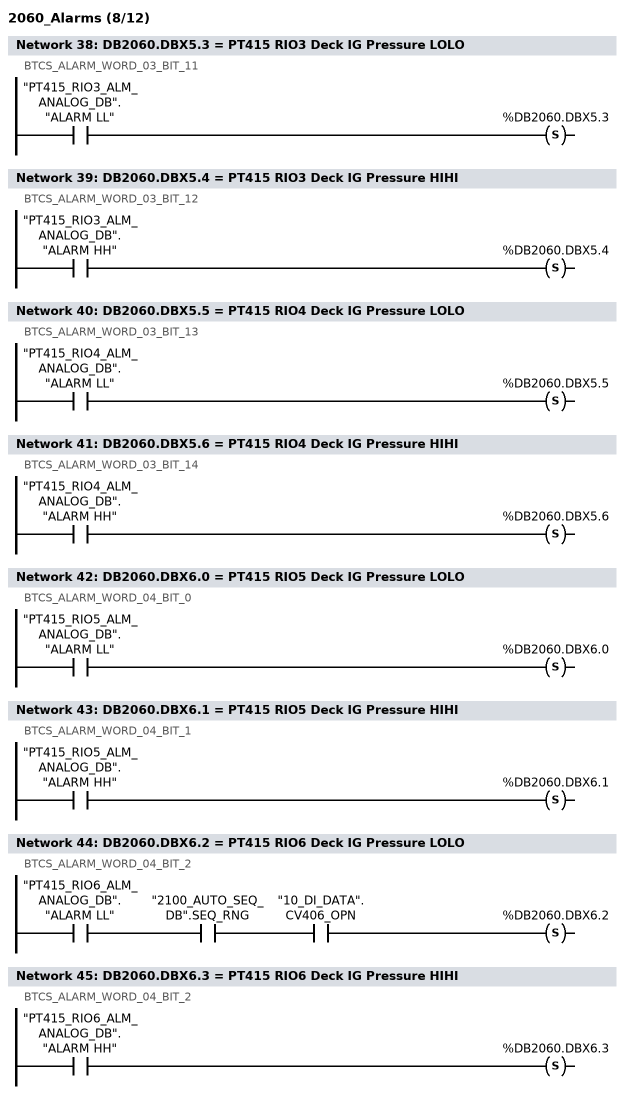
   RUNG wire#powerrail
      Contact( "PT415_RIO3_ALM_ANALOG_DB"."ALARM LL" )
      S_Coil( %DB2060.DBX5.3 )
   END_RUNG
   // the same network as SCL:
   IF "PT415_RIO3_ALM_ANALOG_DB"."ALARM LL" THEN %DB2060.DBX5.3 := TRUE; END_IF;
END_REGION

REGION Network 39: DB2060.DBX5.4 = PT415 RIO3 Deck IG Pressure HIHI
   // BTCS_ALARM_WORD_03_BIT_12
   RUNG wire#powerrail
      Contact( "PT415_RIO3_ALM_ANALOG_DB"."ALARM HH" )
      S_Coil( %DB2060.DBX5.4 )
   END_RUNG
   // the same network as SCL:
   IF "PT415_RIO3_ALM_ANALOG_DB"."ALARM HH" THEN %DB2060.DBX5.4 := TRUE; END_IF;
END_REGION

REGION Network 40: DB2060.DBX5.5 = PT415 RIO4 Deck IG Pressure LOLO
   // BTCS_ALARM_WORD_03_BIT_13
   RUNG wire#powerrail
      Contact( "PT415_RIO4_ALM_ANALOG_DB"."ALARM LL" )
      S_Coil( %DB2060.DBX5.5 )
   END_RUNG
   // the same network as SCL:
   IF "PT415_RIO4_ALM_ANALOG_DB"."ALARM LL" THEN %DB2060.DBX5.5 := TRUE; END_IF;
END_REGION

REGION Network 41: DB2060.DBX5.6 = PT415 RIO4 Deck IG Pressure HIHI
   // BTCS_ALARM_WORD_03_BIT_14
   RUNG wire#powerrail
      Contact( "PT415_RIO4_ALM_ANALOG_DB"."ALARM HH" )
      S_Coil( %DB2060.DBX5.6 )
   END_RUNG
   // the same network as SCL:
   IF "PT415_RIO4_ALM_ANALOG_DB"."ALARM HH" THEN %DB2060.DBX5.6 := TRUE; END_IF;
END_REGION

REGION Network 42: DB2060.DBX6.0 = PT415 RIO5 Deck IG Pressure LOLO
   // BTCS_ALARM_WORD_04_BIT_0
   RUNG wire#powerrail
      Contact( "PT415_RIO5_ALM_ANALOG_DB"."ALARM LL" )
      S_Coil( %DB2060.DBX6.0 )
   END_RUNG
   // the same network as SCL:
   IF "PT415_RIO5_ALM_ANALOG_DB"."ALARM LL" THEN %DB2060.DBX6.0 := TRUE; END_IF;
END_REGION

REGION Network 43: DB2060.DBX6.1 = PT415 RIO5 Deck IG Pressure HIHI
   // BTCS_ALARM_WORD_04_BIT_1
   RUNG wire#powerrail
      Contact( "PT415_RIO5_ALM_ANALOG_DB"."ALARM HH" )
      S_Coil( %DB2060.DBX6.1 )
   END_RUNG
   // the same network as SCL:
   IF "PT415_RIO5_ALM_ANALOG_DB"."ALARM HH" THEN %DB2060.DBX6.1 := TRUE; END_IF;
END_REGION

REGION Network 44: DB2060.DBX6.2 = PT415 RIO6 Deck IG Pressure LOLO
   // BTCS_ALARM_WORD_04_BIT_2
   RUNG wire#powerrail
      Contact( "PT415_RIO6_ALM_ANALOG_DB"."ALARM LL" )
      Contact( "2100_AUTO_SEQ_DB".SEQ_RNG )
      Contact( "10_DI_DATA".CV406_OPN )
      S_Coil( %DB2060.DBX6.2 )
   END_RUNG
   // the same network as SCL:
   IF "PT415_RIO6_ALM_ANALOG_DB"."ALARM LL" AND "2100_AUTO_SEQ_DB".SEQ_RNG AND "10_DI_DATA".CV406_OPN THEN
       %DB2060.DBX6.2 := TRUE;
   END_IF;
END_REGION

REGION Network 45: DB2060.DBX6.3 = PT415 RIO6 Deck IG Pressure HIHI
   // BTCS_ALARM_WORD_04_BIT_2
   RUNG wire#powerrail
      Contact( "PT415_RIO6_ALM_ANALOG_DB"."ALARM HH" )
      S_Coil( %DB2060.DBX6.3 )
   END_RUNG
   // the same network as SCL:
   IF "PT415_RIO6_ALM_ANALOG_DB"."ALARM HH" THEN %DB2060.DBX6.3 := TRUE; END_IF;
END_REGION

REGION Network 46: DB2060.DBX6.4 = PT415 RIO7 Deck IG Pressure LOLO
   // BTCS_ALARM_WORD_04_BIT_4
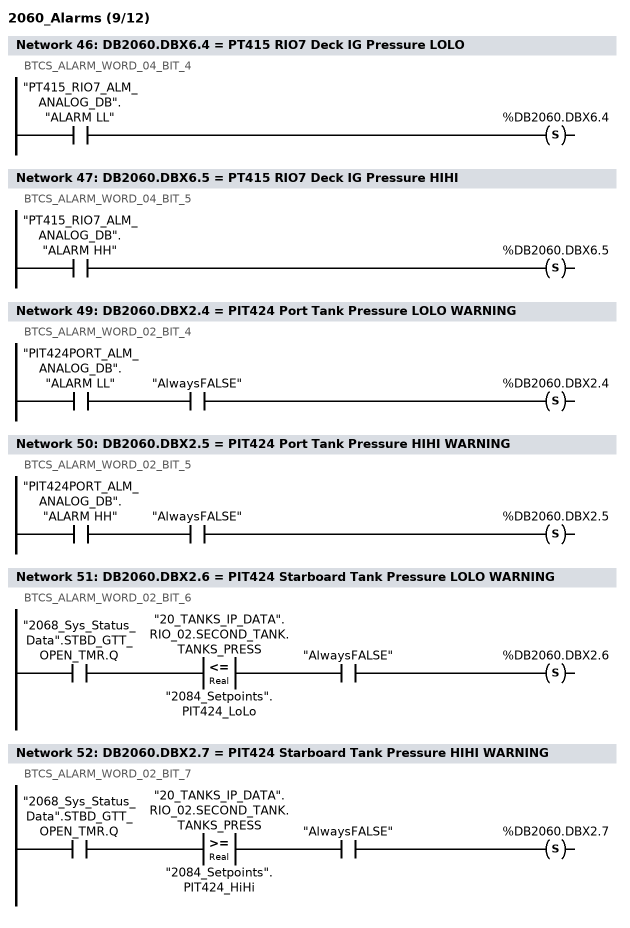
   RUNG wire#powerrail
      Contact( "PT415_RIO7_ALM_ANALOG_DB"."ALARM LL" )
      S_Coil( %DB2060.DBX6.4 )
   END_RUNG
   // the same network as SCL:
   IF "PT415_RIO7_ALM_ANALOG_DB"."ALARM LL" THEN %DB2060.DBX6.4 := TRUE; END_IF;
END_REGION

REGION Network 47: DB2060.DBX6.5 = PT415 RIO7 Deck IG Pressure HIHI
   // BTCS_ALARM_WORD_04_BIT_5
   RUNG wire#powerrail
      Contact( "PT415_RIO7_ALM_ANALOG_DB"."ALARM HH" )
      S_Coil( %DB2060.DBX6.5 )
   END_RUNG
   // the same network as SCL:
   IF "PT415_RIO7_ALM_ANALOG_DB"."ALARM HH" THEN %DB2060.DBX6.5 := TRUE; END_IF;
END_REGION

REGION Network 49: DB2060.DBX2.4 = PIT424 Port Tank Pressure LOLO WARNING
   // BTCS_ALARM_WORD_02_BIT_4
   RUNG wire#powerrail
      Contact( "PIT424PORT_ALM_ANALOG_DB"."ALARM LL" )
      Contact( "AlwaysFALSE" )
      S_Coil( %DB2060.DBX2.4 )
   END_RUNG
   // the same network as SCL:
   IF "PIT424PORT_ALM_ANALOG_DB"."ALARM LL" AND "AlwaysFALSE" THEN %DB2060.DBX2.4 := TRUE; END_IF;
END_REGION

REGION Network 50: DB2060.DBX2.5 = PIT424 Port Tank Pressure HIHI WARNING
   // BTCS_ALARM_WORD_02_BIT_5
   RUNG wire#powerrail
      Contact( "PIT424PORT_ALM_ANALOG_DB"."ALARM HH" )
      Contact( "AlwaysFALSE" )
      S_Coil( %DB2060.DBX2.5 )
   END_RUNG
   // the same network as SCL:
   IF "PIT424PORT_ALM_ANALOG_DB"."ALARM HH" AND "AlwaysFALSE" THEN %DB2060.DBX2.5 := TRUE; END_IF;
END_REGION

REGION Network 51: DB2060.DBX2.6 = PIT424 Starboard Tank Pressure LOLO WARNING
   // BTCS_ALARM_WORD_02_BIT_6
   RUNG wire#powerrail
      Contact( "2068_Sys_Status_Data".STBD_GTT_OPEN_TMR.Q )
      { S7_Templates := "SrcType := Real" } LE_Contact(in1 := "20_TANKS_IP_DATA".RIO_02.SECOND_TANK.TANKS_PRESS, in2 := "2084_Setpoints".PIT424_LoLo)
      Contact( "AlwaysFALSE" )
      S_Coil( %DB2060.DBX2.6 )
   END_RUNG
   // the same network as SCL:
   IF "2068_Sys_Status_Data".STBD_GTT_OPEN_TMR.Q AND ("20_TANKS_IP_DATA".RIO_02.SECOND_TANK.TANKS_PRESS <= "2084_Setpoints".PIT424_LoLo) AND "AlwaysFALSE" THEN
       %DB2060.DBX2.6 := TRUE;
   END_IF;
END_REGION

REGION Network 52: DB2060.DBX2.7 = PIT424 Starboard Tank Pressure HIHI WARNING
   // BTCS_ALARM_WORD_02_BIT_7
   RUNG wire#powerrail
      Contact( "2068_Sys_Status_Data".STBD_GTT_OPEN_TMR.Q )
      { S7_Templates := "SrcType := Real" } GE_Contact(in1 := "20_TANKS_IP_DATA".RIO_02.SECOND_TANK.TANKS_PRESS, in2 := "2084_Setpoints".PIT424_HiHi)
      Contact( "AlwaysFALSE" )
      S_Coil( %DB2060.DBX2.7 )
   END_RUNG
   // the same network as SCL:
   IF "2068_Sys_Status_Data".STBD_GTT_OPEN_TMR.Q AND ("20_TANKS_IP_DATA".RIO_02.SECOND_TANK.TANKS_PRESS >= "2084_Setpoints".PIT424_HiHi) AND "AlwaysFALSE" THEN
       %DB2060.DBX2.7 := TRUE;
   END_IF;
END_REGION

REGION Network 54: Alarm reset
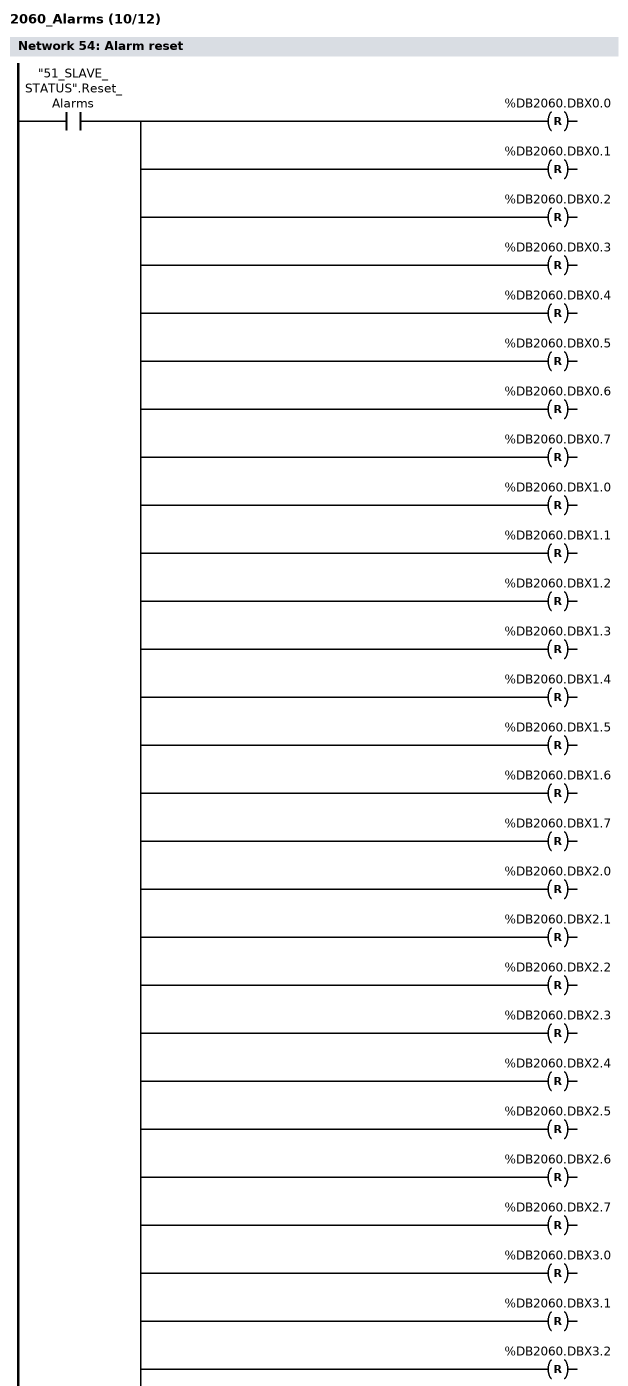
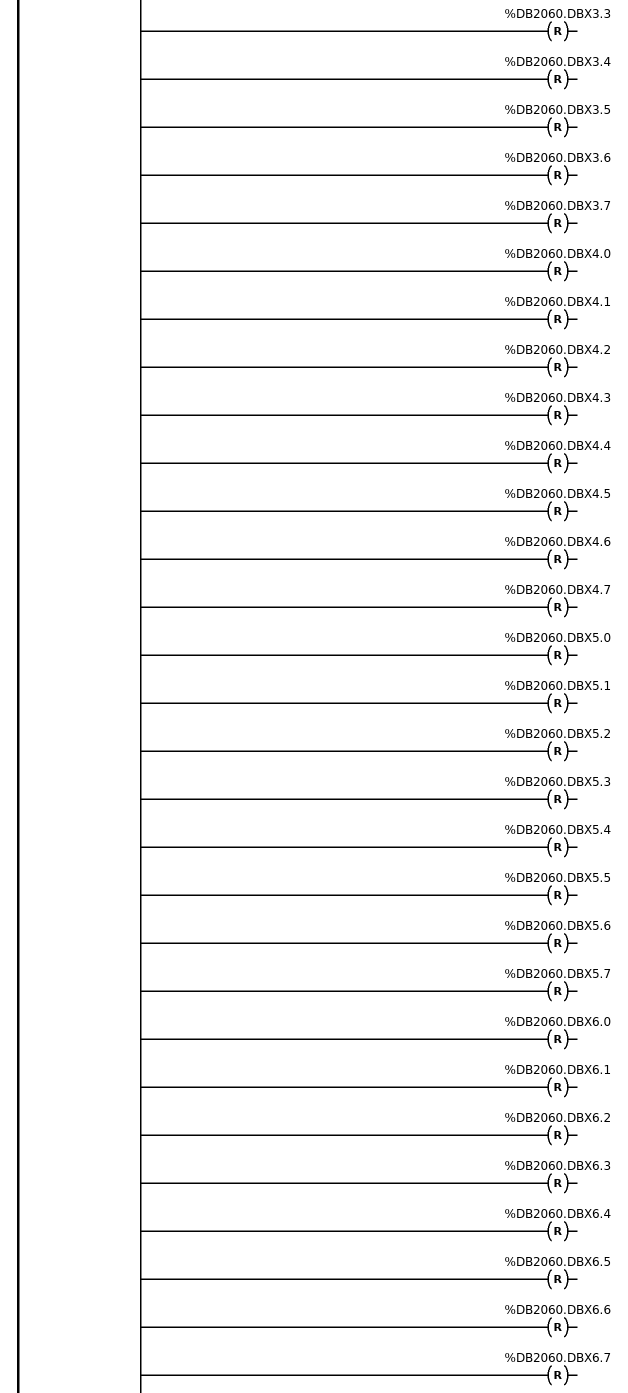
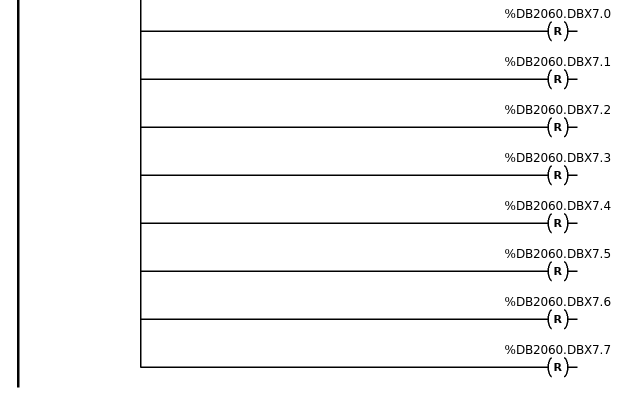
   RUNG wire#powerrail
      Contact( "51_SLAVE_STATUS".Reset_Alarms )
      wire#w1
      R_Coil( %DB2060.DBX0.0 )
   END_RUNG
   RUNG wire#w1
      R_Coil( %DB2060.DBX0.1 )
   END_RUNG
   RUNG wire#w1
      R_Coil( %DB2060.DBX0.2 )
   END_RUNG
   RUNG wire#w1
      R_Coil( %DB2060.DBX0.3 )
   END_RUNG
   RUNG wire#w1
      R_Coil( %DB2060.DBX0.4 )
   END_RUNG
   RUNG wire#w1
      R_Coil( %DB2060.DBX0.5 )
   END_RUNG
   RUNG wire#w1
      R_Coil( %DB2060.DBX0.6 )
   END_RUNG
   RUNG wire#w1
      R_Coil( %DB2060.DBX0.7 )
   END_RUNG
   RUNG wire#w1
      R_Coil( %DB2060.DBX1.0 )
   END_RUNG
   RUNG wire#w1
      R_Coil( %DB2060.DBX1.1 )
   END_RUNG
   RUNG wire#w1
      R_Coil( %DB2060.DBX1.2 )
   END_RUNG
   RUNG wire#w1
      R_Coil( %DB2060.DBX1.3 )
   END_RUNG
   RUNG wire#w1
      R_Coil( %DB2060.DBX1.4 )
   END_RUNG
   RUNG wire#w1
      R_Coil( %DB2060.DBX1.5 )
   END_RUNG
   RUNG wire#w1
      R_Coil( %DB2060.DBX1.6 )
   END_RUNG
   RUNG wire#w1
      R_Coil( %DB2060.DBX1.7 )
   END_RUNG
   RUNG wire#w1
      R_Coil( %DB2060.DBX2.0 )
   END_RUNG
   RUNG wire#w1
      R_Coil( %DB2060.DBX2.1 )
   END_RUNG
   RUNG wire#w1
      R_Coil( %DB2060.DBX2.2 )
   END_RUNG
   RUNG wire#w1
      R_Coil( %DB2060.DBX2.3 )
   END_RUNG
   RUNG wire#w1
      R_Coil( %DB2060.DBX2.4 )
   END_RUNG
   RUNG wire#w1
      R_Coil( %DB2060.DBX2.5 )
   END_RUNG
   RUNG wire#w1
      R_Coil( %DB2060.DBX2.6 )
   END_RUNG
   RUNG wire#w1
      R_Coil( %DB2060.DBX2.7 )
   END_RUNG
   RUNG wire#w1
      R_Coil( %DB2060.DBX3.0 )
   END_RUNG
   RUNG wire#w1
      R_Coil( %DB2060.DBX3.1 )
   END_RUNG
   RUNG wire#w1
      R_Coil( %DB2060.DBX3.2 )
   END_RUNG
   RUNG wire#w1
      R_Coil( %DB2060.DBX3.3 )
   END_RUNG
   RUNG wire#w1
      R_Coil( %DB2060.DBX3.4 )
   END_RUNG
   RUNG wire#w1
      R_Coil( %DB2060.DBX3.5 )
   END_RUNG
   RUNG wire#w1
      R_Coil( %DB2060.DBX3.6 )
   END_RUNG
   RUNG wire#w1
      R_Coil( %DB2060.DBX3.7 )
   END_RUNG
   RUNG wire#w1
      R_Coil( %DB2060.DBX4.0 )
   END_RUNG
   RUNG wire#w1
      R_Coil( %DB2060.DBX4.1 )
   END_RUNG
   RUNG wire#w1
      R_Coil( %DB2060.DBX4.2 )
   END_RUNG
   RUNG wire#w1
      R_Coil( %DB2060.DBX4.3 )
   END_RUNG
   RUNG wire#w1
      R_Coil( %DB2060.DBX4.4 )
   END_RUNG
   RUNG wire#w1
      R_Coil( %DB2060.DBX4.5 )
   END_RUNG
   RUNG wire#w1
      R_Coil( %DB2060.DBX4.6 )
   END_RUNG
   RUNG wire#w1
      R_Coil( %DB2060.DBX4.7 )
   END_RUNG
   RUNG wire#w1
      R_Coil( %DB2060.DBX5.0 )
   END_RUNG
   RUNG wire#w1
      R_Coil( %DB2060.DBX5.1 )
   END_RUNG
   RUNG wire#w1
      R_Coil( %DB2060.DBX5.2 )
   END_RUNG
   RUNG wire#w1
      R_Coil( %DB2060.DBX5.3 )
   END_RUNG
   RUNG wire#w1
      R_Coil( %DB2060.DBX5.4 )
   END_RUNG
   RUNG wire#w1
      R_Coil( %DB2060.DBX5.5 )
   END_RUNG
   RUNG wire#w1
      R_Coil( %DB2060.DBX5.6 )
   END_RUNG
   RUNG wire#w1
      R_Coil( %DB2060.DBX5.7 )
   END_RUNG
   RUNG wire#w1
      R_Coil( %DB2060.DBX6.0 )
   END_RUNG
   RUNG wire#w1
      R_Coil( %DB2060.DBX6.1 )
   END_RUNG
   RUNG wire#w1
      R_Coil( %DB2060.DBX6.2 )
   END_RUNG
   RUNG wire#w1
      R_Coil( %DB2060.DBX6.3 )
   END_RUNG
   RUNG wire#w1
      R_Coil( %DB2060.DBX6.4 )
   END_RUNG
   RUNG wire#w1
      R_Coil( %DB2060.DBX6.5 )
   END_RUNG
   RUNG wire#w1
      R_Coil( %DB2060.DBX6.6 )
   END_RUNG
   RUNG wire#w1
      R_Coil( %DB2060.DBX6.7 )
   END_RUNG
   RUNG wire#w1
      R_Coil( %DB2060.DBX7.0 )
   END_RUNG
   RUNG wire#w1
      R_Coil( %DB2060.DBX7.1 )
   END_RUNG
   RUNG wire#w1
      R_Coil( %DB2060.DBX7.2 )
   END_RUNG
   RUNG wire#w1
      R_Coil( %DB2060.DBX7.3 )
   END_RUNG
   RUNG wire#w1
      R_Coil( %DB2060.DBX7.4 )
   END_RUNG
   RUNG wire#w1
      R_Coil( %DB2060.DBX7.5 )
   END_RUNG
   RUNG wire#w1
      R_Coil( %DB2060.DBX7.6 )
   END_RUNG
   RUNG wire#w1
      R_Coil( %DB2060.DBX7.7 )
   END_RUNG
   // the same network as SCL:
   IF "51_SLAVE_STATUS".Reset_Alarms THEN
       %DB2060.DBX0.0 := FALSE;
       %DB2060.DBX0.1 := FALSE;
       %DB2060.DBX0.2 := FALSE;
       %DB2060.DBX0.3 := FALSE;
       %DB2060.DBX0.4 := FALSE;
       %DB2060.DBX0.5 := FALSE;
       %DB2060.DBX0.6 := FALSE;
       %DB2060.DBX0.7 := FALSE;
       %DB2060.DBX1.0 := FALSE;
       %DB2060.DBX1.1 := FALSE;
       %DB2060.DBX1.2 := FALSE;
       %DB2060.DBX1.3 := FALSE;
       %DB2060.DBX1.4 := FALSE;
       %DB2060.DBX1.5 := FALSE;
       %DB2060.DBX1.6 := FALSE;
       %DB2060.DBX1.7 := FALSE;
       %DB2060.DBX2.0 := FALSE;
       %DB2060.DBX2.1 := FALSE;
       %DB2060.DBX2.2 := FALSE;
       %DB2060.DBX2.3 := FALSE;
       %DB2060.DBX2.4 := FALSE;
       %DB2060.DBX2.5 := FALSE;
       %DB2060.DBX2.6 := FALSE;
       %DB2060.DBX2.7 := FALSE;
       %DB2060.DBX3.0 := FALSE;
       %DB2060.DBX3.1 := FALSE;
       %DB2060.DBX3.2 := FALSE;
       %DB2060.DBX3.3 := FALSE;
       %DB2060.DBX3.4 := FALSE;
       %DB2060.DBX3.5 := FALSE;
       %DB2060.DBX3.6 := FALSE;
       %DB2060.DBX3.7 := FALSE;
       %DB2060.DBX4.0 := FALSE;
       %DB2060.DBX4.1 := FALSE;
       %DB2060.DBX4.2 := FALSE;
       %DB2060.DBX4.3 := FALSE;
       %DB2060.DBX4.4 := FALSE;
       %DB2060.DBX4.5 := FALSE;
       %DB2060.DBX4.6 := FALSE;
       %DB2060.DBX4.7 := FALSE;
       %DB2060.DBX5.0 := FALSE;
       %DB2060.DBX5.1 := FALSE;
       %DB2060.DBX5.2 := FALSE;
       %DB2060.DBX5.3 := FALSE;
       %DB2060.DBX5.4 := FALSE;
       %DB2060.DBX5.5 := FALSE;
       %DB2060.DBX5.6 := FALSE;
       %DB2060.DBX5.7 := FALSE;
       %DB2060.DBX6.0 := FALSE;
       %DB2060.DBX6.1 := FALSE;
       %DB2060.DBX6.2 := FALSE;
       %DB2060.DBX6.3 := FALSE;
       %DB2060.DBX6.4 := FALSE;
       %DB2060.DBX6.5 := FALSE;
       %DB2060.DBX6.6 := FALSE;
       %DB2060.DBX6.7 := FALSE;
       %DB2060.DBX7.0 := FALSE;
       %DB2060.DBX7.1 := FALSE;
       %DB2060.DBX7.2 := FALSE;
       %DB2060.DBX7.3 := FALSE;
       %DB2060.DBX7.4 := FALSE;
       %DB2060.DBX7.5 := FALSE;
       %DB2060.DBX7.6 := FALSE;
       %DB2060.DBX7.7 := FALSE;
   END_IF;
END_REGION

REGION Network 55: New Alarm
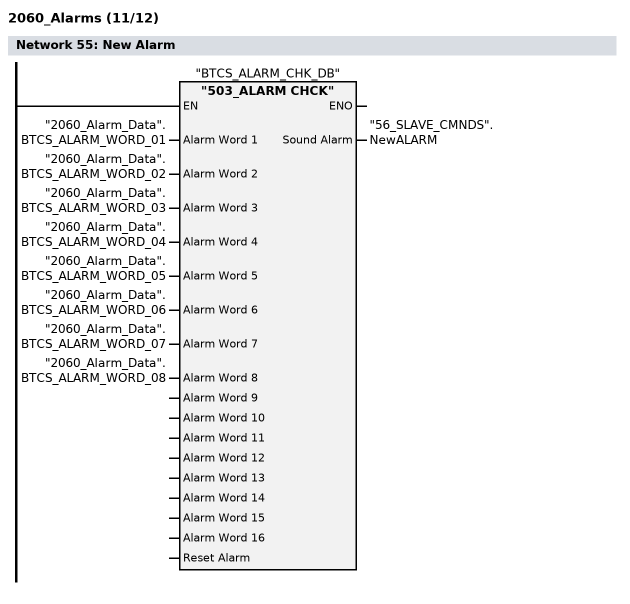
   RUNG wire#powerrail
      "BTCS_ALARM_CHK_DB"("Alarm Word 1" := "2060_Alarm_Data".BTCS_ALARM_WORD_01, "Alarm Word 2" := "2060_Alarm_Data".BTCS_ALARM_WORD_02, "Alarm Word 3" := "2060_Alarm_Data".BTCS_ALARM_WORD_03, "Alarm Word 4" := "2060_Alarm_Data".BTCS_ALARM_WORD_04, "Alarm Word 5" := "2060_Alarm_Data".BTCS_ALARM_WORD_05, "Alarm Word 6" := "2060_Alarm_Data".BTCS_ALARM_WORD_06, "Alarm Word 7" := "2060_Alarm_Data".BTCS_ALARM_WORD_07, "Alarm Word 8" := "2060_Alarm_Data".BTCS_ALARM_WORD_08, "Alarm Word 9" :=, "Alarm Word 10" :=, "Alarm Word 11" :=, "Alarm Word 12" :=, "Alarm Word 13" :=, "Alarm Word 14" :=, "Alarm Word 15" :=, "Alarm Word 16" :=, "Reset Alarm" :=, "Sound Alarm" => "56_SLAVE_CMNDS".NewALARM)
   END_RUNG
   // the same network as SCL:
   "BTCS_ALARM_CHK_DB"("Alarm Word 1" := "2060_Alarm_Data".BTCS_ALARM_WORD_01,   // "503_ALARM CHCK"
                       "Alarm Word 2" := "2060_Alarm_Data".BTCS_ALARM_WORD_02,
                       "Alarm Word 3" := "2060_Alarm_Data".BTCS_ALARM_WORD_03,
                       "Alarm Word 4" := "2060_Alarm_Data".BTCS_ALARM_WORD_04,
                       "Alarm Word 5" := "2060_Alarm_Data".BTCS_ALARM_WORD_05,
                       "Alarm Word 6" := "2060_Alarm_Data".BTCS_ALARM_WORD_06,
                       "Alarm Word 7" := "2060_Alarm_Data".BTCS_ALARM_WORD_07,
                       "Alarm Word 8" := "2060_Alarm_Data".BTCS_ALARM_WORD_08,
                       "Sound Alarm" => "56_SLAVE_CMNDS".NewALARM);
END_REGION

REGION Network 56: Alarm Present
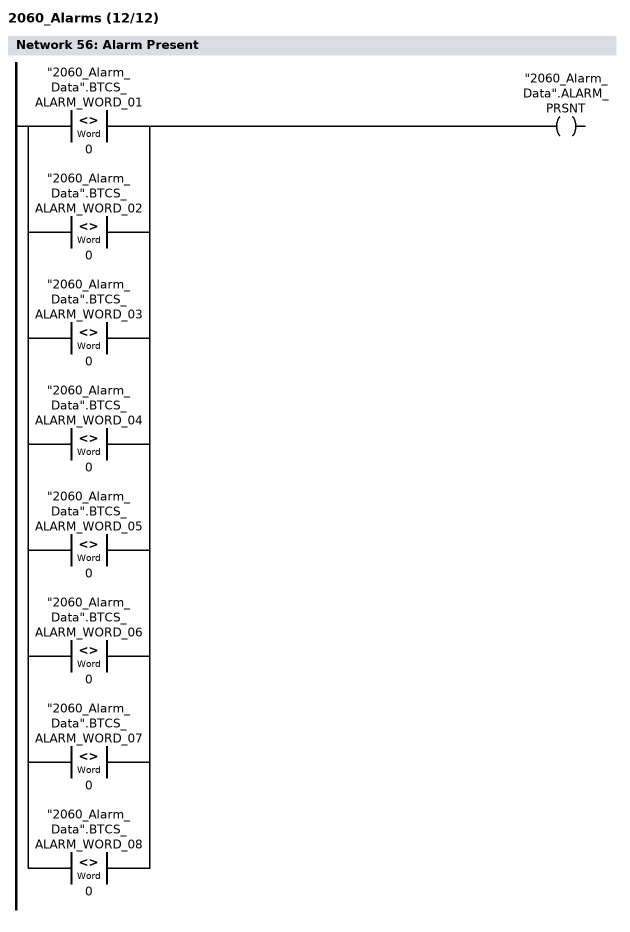
   RUNG wire#powerrail
      { S7_Templates := "SrcType := Word" } NE_Contact(in1 := "2060_Alarm_Data".BTCS_ALARM_WORD_01, in2 := 0)
      wire#w1
      Coil( "2060_Alarm_Data".ALARM_PRSNT )
   END_RUNG
   RUNG wire#powerrail
      { S7_Templates := "SrcType := Word" } NE_Contact(in1 := "2060_Alarm_Data".BTCS_ALARM_WORD_02, in2 := 0)
   END_RUNG wire#w1
   RUNG wire#powerrail
      { S7_Templates := "SrcType := Word" } NE_Contact(in1 := "2060_Alarm_Data".BTCS_ALARM_WORD_03, in2 := 0)
   END_RUNG wire#w1
   RUNG wire#powerrail
      { S7_Templates := "SrcType := Word" } NE_Contact(in1 := "2060_Alarm_Data".BTCS_ALARM_WORD_04, in2 := 0)
   END_RUNG wire#w1
   RUNG wire#powerrail
      { S7_Templates := "SrcType := Word" } NE_Contact(in1 := "2060_Alarm_Data".BTCS_ALARM_WORD_05, in2 := 0)
   END_RUNG wire#w1
   RUNG wire#powerrail
      { S7_Templates := "SrcType := Word" } NE_Contact(in1 := "2060_Alarm_Data".BTCS_ALARM_WORD_06, in2 := 0)
   END_RUNG wire#w1
   RUNG wire#powerrail
      { S7_Templates := "SrcType := Word" } NE_Contact(in1 := "2060_Alarm_Data".BTCS_ALARM_WORD_07, in2 := 0)
   END_RUNG wire#w1
   RUNG wire#powerrail
      { S7_Templates := "SrcType := Word" } NE_Contact(in1 := "2060_Alarm_Data".BTCS_ALARM_WORD_08, in2 := 0)
   END_RUNG wire#w1
   // the same network as SCL:
   "2060_Alarm_Data".ALARM_PRSNT := ("2060_Alarm_Data".BTCS_ALARM_WORD_01 <> 0) OR ("2060_Alarm_Data".BTCS_ALARM_WORD_02 <> 0) OR ("2060_Alarm_Data".BTCS_ALARM_WORD_03 <> 0) OR ("2060_Alarm_Data".BTCS_ALARM_WORD_04 <> 0) OR ("2060_Alarm_Data".BTCS_ALARM_WORD_05 <> 0) OR ("2060_Alarm_Data".BTCS_ALARM_WORD_06 <> 0) OR ("2060_Alarm_Data".BTCS_ALARM_WORD_07 <> 0) OR ("2060_Alarm_Data".BTCS_ALARM_WORD_08 <> 0);
END_REGION
END_FUNCTION

FUNCTION "2062_Warnings" : Void   // FC2062, LAD
TITLE = Warning Processing
{ S7_Optimized_Access := 'TRUE' }
AUTHOR : JRS
VERSION : 0.1
// To warning conditions
   VAR_TEMP   // added for the SCL form of the ladder/FBD networks
      _w1 : Bool;
   END_VAR
BEGIN

REGION Network 1: DB2062 DBX0.0 = 600-TX-433 RIO7 Confined Space O2 Monitor
   // BTCS_WARNING_WORD_01_BIT_0                           15.10
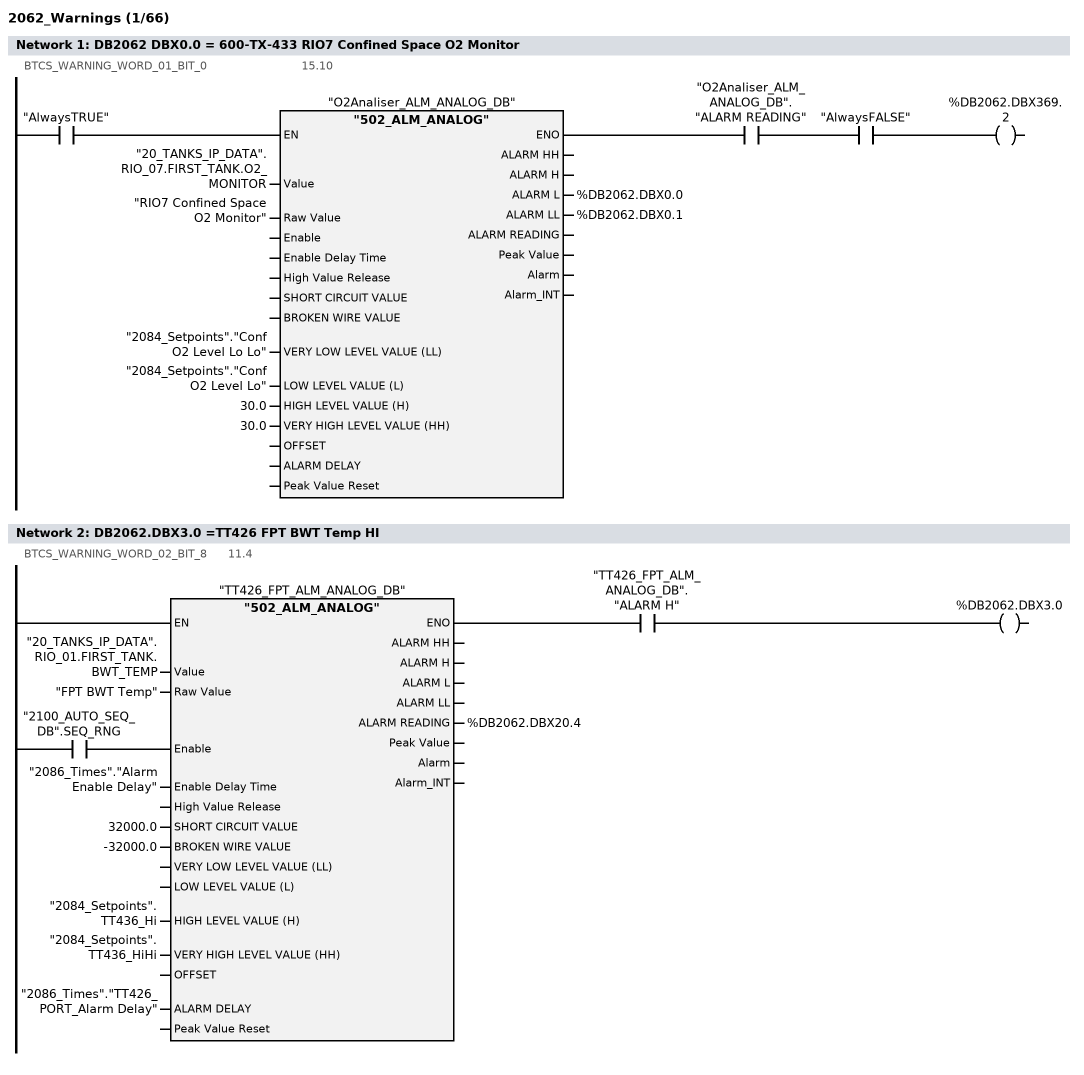
   RUNG wire#powerrail
      Contact( "AlwaysTRUE" )
      "O2Analiser_ALM_ANALOG_DB"(Value := "20_TANKS_IP_DATA".RIO_07.FIRST_TANK.O2_MONITOR, "Raw Value" := "RIO7 Confined Space O2 Monitor", Enable :=, "Enable Delay Time" :=, "High Value Release" :=, "SHORT CIRCUIT VALUE" :=, "BROKEN WIRE VALUE" :=, "VERY LOW LEVEL VALUE (LL)" := "2084_Setpoints"."Conf O2 Level Lo Lo", "LOW LEVEL VALUE (L)" := "2084_Setpoints"."Conf O2 Level Lo", "HIGH LEVEL VALUE (H)" := 30.0, "VERY HIGH LEVEL VALUE (HH)" := 30.0, OFFSET :=, "ALARM DELAY" :=, "Peak Value Reset" :=, "ALARM HH" =>, "ALARM H" =>, "ALARM L" => %DB2062.DBX0.0, "ALARM LL" => %DB2062.DBX0.1, "ALARM READING" =>, "Peak Value" =>, Alarm =>, Alarm_INT =>)
      Contact( "O2Analiser_ALM_ANALOG_DB"."ALARM READING" )
      Contact( "AlwaysFALSE" )
      Coil( %DB2062.DBX369.2 )
   END_RUNG
   // the same network as SCL:
   "O2Analiser_ALM_ANALOG_DB"(EN := "AlwaysTRUE",   // "502_ALM_ANALOG"
                           Value := "20_TANKS_IP_DATA".RIO_07.FIRST_TANK.O2_MONITOR,
                           "Raw Value" := "RIO7 Confined Space O2 Monitor",
                           "VERY LOW LEVEL VALUE (LL)" := "2084_Setpoints"."Conf O2 Level Lo Lo",
                           "LOW LEVEL VALUE (L)" := "2084_Setpoints"."Conf O2 Level Lo",
                           "HIGH LEVEL VALUE (H)" := 30.0,
                           "VERY HIGH LEVEL VALUE (HH)" := 30.0,
                           "ALARM L" => %DB2062.DBX0.0,
                           "ALARM LL" => %DB2062.DBX0.1,
                           ENO => #_w1);
   %DB2062.DBX369.2 := #_w1 AND "O2Analiser_ALM_ANALOG_DB"."ALARM READING" AND "AlwaysFALSE";
END_REGION

REGION Network 2: DB2062.DBX3.0 =TT426 FPT BWT Temp HI
   // BTCS_WARNING_WORD_02_BIT_8      11.4
   RUNG wire#powerrail
      "TT426_FPT_ALM_ANALOG_DB"(Enable := wire#w1, Value := "20_TANKS_IP_DATA".RIO_01.FIRST_TANK.BWT_TEMP, "Raw Value" := "FPT BWT Temp", "Enable Delay Time" := "2086_Times"."Alarm Enable Delay", "High Value Release" :=, "SHORT CIRCUIT VALUE" := 32000.0, "BROKEN WIRE VALUE" := -32000.0, "VERY LOW LEVEL VALUE (LL)" :=, "LOW LEVEL VALUE (L)" :=, "HIGH LEVEL VALUE (H)" := "2084_Setpoints".TT436_Hi, "VERY HIGH LEVEL VALUE (HH)" := "2084_Setpoints".TT436_HiHi, OFFSET :=, "ALARM DELAY" := "2086_Times"."TT426_PORT_Alarm Delay", "Peak Value Reset" :=, "ALARM HH" =>, "ALARM H" =>, "ALARM L" =>, "ALARM LL" =>, "ALARM READING" => %DB2062.DBX20.4, "Peak Value" =>, Alarm =>, Alarm_INT =>)
      Contact( "TT426_FPT_ALM_ANALOG_DB"."ALARM H" )
      Coil( %DB2062.DBX3.0 )
   END_RUNG
   RUNG wire#powerrail
      Contact( "2100_AUTO_SEQ_DB".SEQ_RNG )
   END_RUNG wire#w1
   // the same network as SCL:
   "TT426_FPT_ALM_ANALOG_DB"(Value := "20_TANKS_IP_DATA".RIO_01.FIRST_TANK.BWT_TEMP,   // "502_ALM_ANALOG"
                           "Raw Value" := "FPT BWT Temp",
                           Enable := "2100_AUTO_SEQ_DB".SEQ_RNG,
                           "Enable Delay Time" := "2086_Times"."Alarm Enable Delay",
                           "SHORT CIRCUIT VALUE" := 32000.0,
                           "BROKEN WIRE VALUE" := -32000.0,
                           "HIGH LEVEL VALUE (H)" := "2084_Setpoints".TT436_Hi,
                           "VERY HIGH LEVEL VALUE (HH)" := "2084_Setpoints".TT436_HiHi,
                           "ALARM DELAY" := "2086_Times"."TT426_PORT_Alarm Delay",
                           "ALARM READING" => %DB2062.DBX20.4,
                           ENO => #_w1);
   %DB2062.DBX3.0 := #_w1 AND "TT426_FPT_ALM_ANALOG_DB"."ALARM H";
END_REGION

REGION Network 3: DB2062.DBX3.1 =TT426 1P BWT Temp HI
   // BTCS_WARNING_WORD_02_BIT_9                   11.5
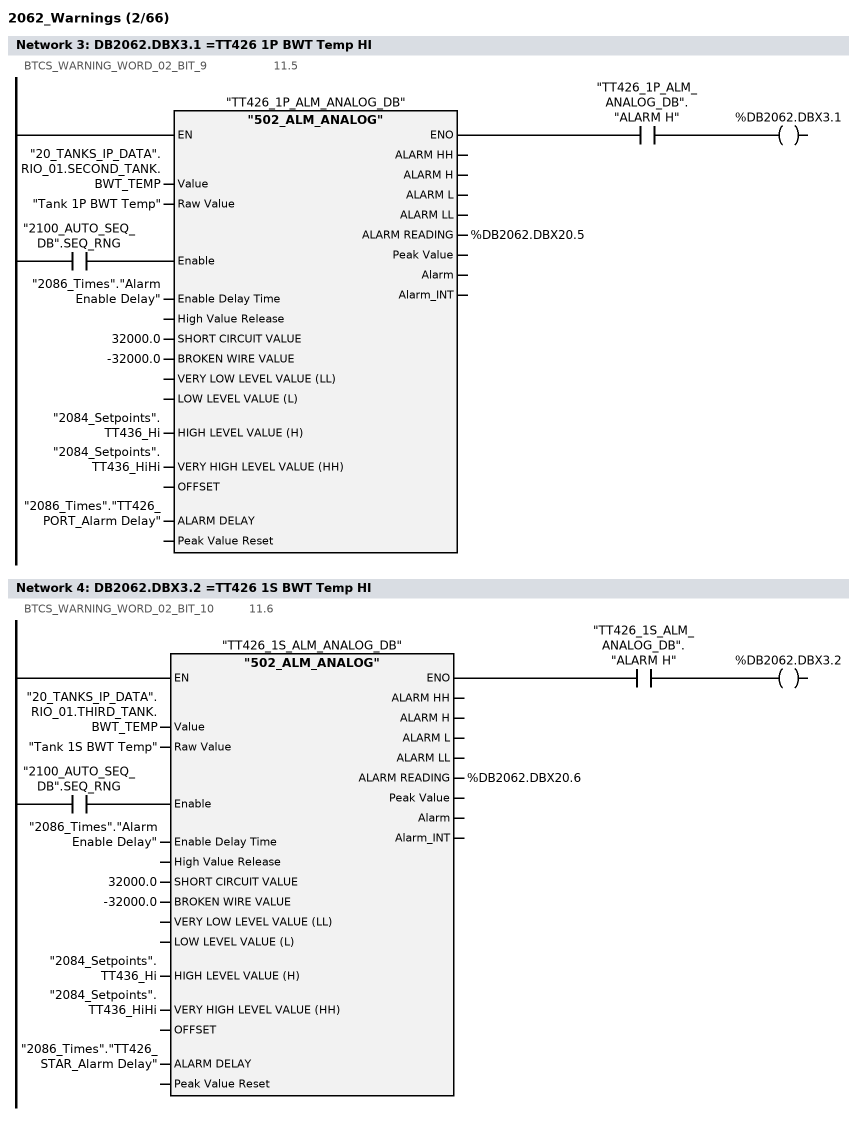
   RUNG wire#powerrail
      "TT426_1P_ALM_ANALOG_DB"(Enable := wire#w1, Value := "20_TANKS_IP_DATA".RIO_01.SECOND_TANK.BWT_TEMP, "Raw Value" := "Tank 1P BWT Temp", "Enable Delay Time" := "2086_Times"."Alarm Enable Delay", "High Value Release" :=, "SHORT CIRCUIT VALUE" := 32000.0, "BROKEN WIRE VALUE" := -32000.0, "VERY LOW LEVEL VALUE (LL)" :=, "LOW LEVEL VALUE (L)" :=, "HIGH LEVEL VALUE (H)" := "2084_Setpoints".TT436_Hi, "VERY HIGH LEVEL VALUE (HH)" := "2084_Setpoints".TT436_HiHi, OFFSET :=, "ALARM DELAY" := "2086_Times"."TT426_PORT_Alarm Delay", "Peak Value Reset" :=, "ALARM HH" =>, "ALARM H" =>, "ALARM L" =>, "ALARM LL" =>, "ALARM READING" => %DB2062.DBX20.5, "Peak Value" =>, Alarm =>, Alarm_INT =>)
      Contact( "TT426_1P_ALM_ANALOG_DB"."ALARM H" )
      Coil( %DB2062.DBX3.1 )
   END_RUNG
   RUNG wire#powerrail
      Contact( "2100_AUTO_SEQ_DB".SEQ_RNG )
   END_RUNG wire#w1
   // the same network as SCL:
   "TT426_1P_ALM_ANALOG_DB"(Value := "20_TANKS_IP_DATA".RIO_01.SECOND_TANK.BWT_TEMP,   // "502_ALM_ANALOG"
                           "Raw Value" := "Tank 1P BWT Temp",
                           Enable := "2100_AUTO_SEQ_DB".SEQ_RNG,
                           "Enable Delay Time" := "2086_Times"."Alarm Enable Delay",
                           "SHORT CIRCUIT VALUE" := 32000.0,
                           "BROKEN WIRE VALUE" := -32000.0,
                           "HIGH LEVEL VALUE (H)" := "2084_Setpoints".TT436_Hi,
                           "VERY HIGH LEVEL VALUE (HH)" := "2084_Setpoints".TT436_HiHi,
                           "ALARM DELAY" := "2086_Times"."TT426_PORT_Alarm Delay",
                           "ALARM READING" => %DB2062.DBX20.5,
                           ENO => #_w1);
   %DB2062.DBX3.1 := #_w1 AND "TT426_1P_ALM_ANALOG_DB"."ALARM H";
END_REGION

REGION Network 4: DB2062.DBX3.2 =TT426 1S BWT Temp HI
   // BTCS_WARNING_WORD_02_BIT_10          11.6
   RUNG wire#powerrail
      "TT426_1S_ALM_ANALOG_DB"(Enable := wire#w1, Value := "20_TANKS_IP_DATA".RIO_01.THIRD_TANK.BWT_TEMP, "Raw Value" := "Tank 1S BWT Temp", "Enable Delay Time" := "2086_Times"."Alarm Enable Delay", "High Value Release" :=, "SHORT CIRCUIT VALUE" := 32000.0, "BROKEN WIRE VALUE" := -32000.0, "VERY LOW LEVEL VALUE (LL)" :=, "LOW LEVEL VALUE (L)" :=, "HIGH LEVEL VALUE (H)" := "2084_Setpoints".TT436_Hi, "VERY HIGH LEVEL VALUE (HH)" := "2084_Setpoints".TT436_HiHi, OFFSET :=, "ALARM DELAY" := "2086_Times"."TT426_STAR_Alarm Delay", "Peak Value Reset" :=, "ALARM HH" =>, "ALARM H" =>, "ALARM L" =>, "ALARM LL" =>, "ALARM READING" => %DB2062.DBX20.6, "Peak Value" =>, Alarm =>, Alarm_INT =>)
      Contact( "TT426_1S_ALM_ANALOG_DB"."ALARM H" )
      Coil( %DB2062.DBX3.2 )
   END_RUNG
   RUNG wire#powerrail
      Contact( "2100_AUTO_SEQ_DB".SEQ_RNG )
   END_RUNG wire#w1
   // the same network as SCL:
   "TT426_1S_ALM_ANALOG_DB"(Value := "20_TANKS_IP_DATA".RIO_01.THIRD_TANK.BWT_TEMP,   // "502_ALM_ANALOG"
                           "Raw Value" := "Tank 1S BWT Temp",
                           Enable := "2100_AUTO_SEQ_DB".SEQ_RNG,
                           "Enable Delay Time" := "2086_Times"."Alarm Enable Delay",
                           "SHORT CIRCUIT VALUE" := 32000.0,
                           "BROKEN WIRE VALUE" := -32000.0,
                           "HIGH LEVEL VALUE (H)" := "2084_Setpoints".TT436_Hi,
                           "VERY HIGH LEVEL VALUE (HH)" := "2084_Setpoints".TT436_HiHi,
                           "ALARM DELAY" := "2086_Times"."TT426_STAR_Alarm Delay",
                           "ALARM READING" => %DB2062.DBX20.6,
                           ENO => #_w1);
   %DB2062.DBX3.2 := #_w1 AND "TT426_1S_ALM_ANALOG_DB"."ALARM H";
END_REGION

REGION Network 5: DB2062.DBX0.2 = TT426 2P BWT Temp HI
   // BTCS_WARNING_WORD_01_BIT_2          11.7
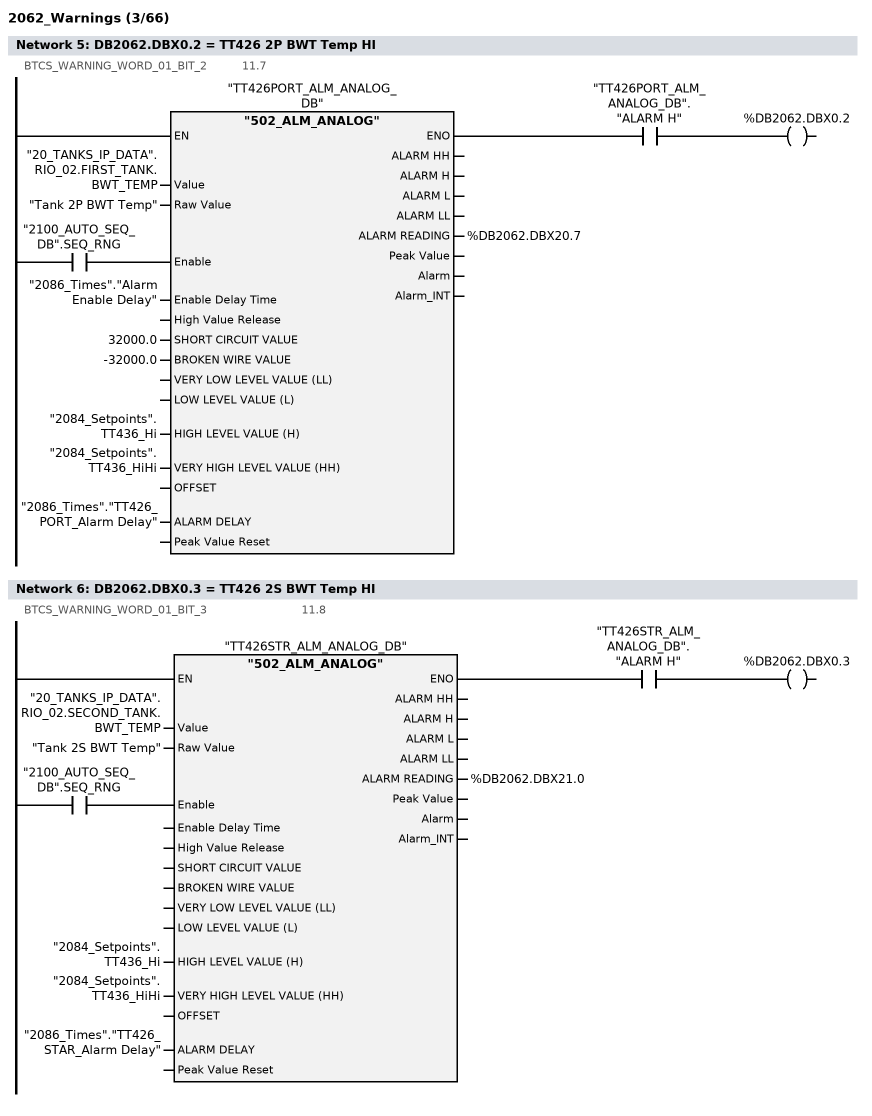
   RUNG wire#powerrail
      "TT426PORT_ALM_ANALOG_DB"(Enable := wire#w1, Value := "20_TANKS_IP_DATA".RIO_02.FIRST_TANK.BWT_TEMP, "Raw Value" := "Tank 2P BWT Temp", "Enable Delay Time" := "2086_Times"."Alarm Enable Delay", "High Value Release" :=, "SHORT CIRCUIT VALUE" := 32000.0, "BROKEN WIRE VALUE" := -32000.0, "VERY LOW LEVEL VALUE (LL)" :=, "LOW LEVEL VALUE (L)" :=, "HIGH LEVEL VALUE (H)" := "2084_Setpoints".TT436_Hi, "VERY HIGH LEVEL VALUE (HH)" := "2084_Setpoints".TT436_HiHi, OFFSET :=, "ALARM DELAY" := "2086_Times"."TT426_PORT_Alarm Delay", "Peak Value Reset" :=, "ALARM HH" =>, "ALARM H" =>, "ALARM L" =>, "ALARM LL" =>, "ALARM READING" => %DB2062.DBX20.7, "Peak Value" =>, Alarm =>, Alarm_INT =>)
      Contact( "TT426PORT_ALM_ANALOG_DB"."ALARM H" )
      Coil( %DB2062.DBX0.2 )
   END_RUNG
   RUNG wire#powerrail
      Contact( "2100_AUTO_SEQ_DB".SEQ_RNG )
   END_RUNG wire#w1
   // the same network as SCL:
   "TT426PORT_ALM_ANALOG_DB"(Value := "20_TANKS_IP_DATA".RIO_02.FIRST_TANK.BWT_TEMP,   // "502_ALM_ANALOG"
                           "Raw Value" := "Tank 2P BWT Temp",
                           Enable := "2100_AUTO_SEQ_DB".SEQ_RNG,
                           "Enable Delay Time" := "2086_Times"."Alarm Enable Delay",
                           "SHORT CIRCUIT VALUE" := 32000.0,
                           "BROKEN WIRE VALUE" := -32000.0,
                           "HIGH LEVEL VALUE (H)" := "2084_Setpoints".TT436_Hi,
                           "VERY HIGH LEVEL VALUE (HH)" := "2084_Setpoints".TT436_HiHi,
                           "ALARM DELAY" := "2086_Times"."TT426_PORT_Alarm Delay",
                           "ALARM READING" => %DB2062.DBX20.7,
                           ENO => #_w1);
   %DB2062.DBX0.2 := #_w1 AND "TT426PORT_ALM_ANALOG_DB"."ALARM H";
END_REGION

REGION Network 6: DB2062.DBX0.3 = TT426 2S BWT Temp HI
   // BTCS_WARNING_WORD_01_BIT_3                           11.8
   RUNG wire#powerrail
      "TT426STR_ALM_ANALOG_DB"(Enable := wire#w1, Value := "20_TANKS_IP_DATA".RIO_02.SECOND_TANK.BWT_TEMP, "Raw Value" := "Tank 2S BWT Temp", "Enable Delay Time" :=, "High Value Release" :=, "SHORT CIRCUIT VALUE" :=, "BROKEN WIRE VALUE" :=, "VERY LOW LEVEL VALUE (LL)" :=, "LOW LEVEL VALUE (L)" :=, "HIGH LEVEL VALUE (H)" := "2084_Setpoints".TT436_Hi, "VERY HIGH LEVEL VALUE (HH)" := "2084_Setpoints".TT436_HiHi, OFFSET :=, "ALARM DELAY" := "2086_Times"."TT426_STAR_Alarm Delay", "Peak Value Reset" :=, "ALARM HH" =>, "ALARM H" =>, "ALARM L" =>, "ALARM LL" =>, "ALARM READING" => %DB2062.DBX21.0, "Peak Value" =>, Alarm =>, Alarm_INT =>)
      Contact( "TT426STR_ALM_ANALOG_DB"."ALARM H" )
      Coil( %DB2062.DBX0.3 )
   END_RUNG
   RUNG wire#powerrail
      Contact( "2100_AUTO_SEQ_DB".SEQ_RNG )
   END_RUNG wire#w1
   // the same network as SCL:
   "TT426STR_ALM_ANALOG_DB"(Value := "20_TANKS_IP_DATA".RIO_02.SECOND_TANK.BWT_TEMP,   // "502_ALM_ANALOG"
                           "Raw Value" := "Tank 2S BWT Temp",
                           Enable := "2100_AUTO_SEQ_DB".SEQ_RNG,
                           "HIGH LEVEL VALUE (H)" := "2084_Setpoints".TT436_Hi,
                           "VERY HIGH LEVEL VALUE (HH)" := "2084_Setpoints".TT436_HiHi,
                           "ALARM DELAY" := "2086_Times"."TT426_STAR_Alarm Delay",
                           "ALARM READING" => %DB2062.DBX21.0,
                           ENO => #_w1);
   %DB2062.DBX0.3 := #_w1 AND "TT426STR_ALM_ANALOG_DB"."ALARM H";
END_REGION

REGION Network 7: DB2062.DBX3.3 =TT426 3P BWT Temp HI
   // BTCS_WARNING_WORD_02_BIT_11                11.9